VERSION : 0.1
   VAR_INPUT
      initValue : DWord;   // Initial value of CRC
      mask : DWord;   // Mask (CRC polynomial) / generator polynomial
      finalXorValue : DWord;   // Value to XOR the result with
      reflectInput : Bool;   // Reflect input (bits are used in reverse order)
      reflectResult : Bool;   // Reflect result (bits are used in reverse order)
   END_VAR
   VAR_IN_OUT
      inputArray : Array[*] of Byte;   // Input array / data stream
   END_VAR
   VAR_TEMP
      tempInput : Byte;   // Current input byte
      tempCRC : DWord;   // CRC checksum
      tempInvCRC : DWord;   // Inverted CRC checksum
      tempLowerLimit : DInt;   // Lower limit of input array
      tempUpperLimit : DInt;   // Upper limit of input array
      tempIndex1 : Int;   // -
      tempIndex2 : Int;   // -
   END_VAR
   // Ret_Val : CRC32 checksum
BEGIN
   //=============================================================================
   // Siemens AG
   // (c)Copyright 2017
   //-----------------------------------------------------------------------------
   // Library:       LGF (Library General Functions)
   // Tested with:   CPU1212C DC/DC/DC FW:V4.2
   // Engineering:   TIA Portal V14 SP1 Upd 5
   // Restrictions:  -
   // Requirements:  PLC (S7-1200 / S7-1500)
   // Functionality: CRC32
   //-----------------------------------------------------------------------------
   // Change log table:
   // Version  Date        In charge / Changes applied
   // 01.00.00 03.07.2018  Siemens Industry Online Support
   //                      First released version
   // 01.00.01 17.08.2018  Siemens Industry Online Support
   //                      Upgrade: TIA V15 Update 2
   // 01.00.02 23.11.2018  Siemens Industry Online Support
   //                      Upgrade: TIA V15.1
   //=============================================================================

   #tempLowerLimit := LOWER_BOUND(ARR := #inputArray, DIM := 1);
   #tempUpperLimit := UPPER_BOUND(ARR := #inputArray, DIM := 1);

   #tempCRC := #initValue;

   FOR #tempIndex1 := #tempLowerLimit TO #tempUpperLimit DO

     IF (#reflectInput = TRUE)
     THEN
       // Reverse bit order in input byte
       #tempInput.%X7 := #inputArray[#tempIndex1].%X0;
       #tempInput.%X6 := #inputArray[#tempIndex1].%X1;
       #tempInput.%X5 := #inputArray[#tempIndex1].%X2;
       #tempInput.%X4 := #inputArray[#tempIndex1].%X3;
       #tempInput.%X3 := #inputArray[#tempIndex1].%X4;
       #tempInput.%X2 := #inputArray[#tempIndex1].%X5;
       #tempInput.%X1 := #inputArray[#tempIndex1].%X6;
       #tempInput.%X0 := #inputArray[#tempIndex1].%X7;
     ELSE
       #tempInput := #inputArray[#tempIndex1];
     END_IF;

     #tempCRC := #tempCRC XOR SHL(IN := BYTE_TO_DWORD(#tempInput), N := 24);

     FOR #tempIndex2 := 0 TO 7 DO
       IF ((#tempCRC AND 16#80000000) <> 0)
       THEN
         #tempCRC := SHL(IN := #tempCRC, N := 1) XOR #mask;
       ELSE
         #tempCRC := SHL(IN := #tempCRC, N := 1);
       END_IF;
     END_FOR;

   END_FOR;

   IF (#reflectResult = TRUE)
   THEN
     // Reverse bit order in CRC checksum
     #tempInvCRC.%X31 := #tempCRC.%X0;
     #tempInvCRC.%X30 := #tempCRC.%X1;
     #tempInvCRC.%X29 := #tempCRC.%X2;
     #tempInvCRC.%X28 := #tempCRC.%X3;
     #tempInvCRC.%X27 := #tempCRC.%X4;
     #tempInvCRC.%X26 := #tempCRC.%X5;
     #tempInvCRC.%X25 := #tempCRC.%X6;
     #tempInvCRC.%X24 := #tempCRC.%X7;
     #tempInvCRC.%X23 := #tempCRC.%X8;
     #tempInvCRC.%X22 := #tempCRC.%X9;
     #tempInvCRC.%X21 := #tempCRC.%X10;
     #tempInvCRC.%X20 := #tempCRC.%X11;
     #tempInvCRC.%X19 := #tempCRC.%X12;
     #tempInvCRC.%X18 := #tempCRC.%X13;
     #tempInvCRC.%X17 := #tempCRC.%X14;
     #tempInvCRC.%X16 := #tempCRC.%X15;
     #tempInvCRC.%X15 := #tempCRC.%X16;
     #tempInvCRC.%X14 := #tempCRC.%X17;
     #tempInvCRC.%X13 := #tempCRC.%X18;
     #tempInvCRC.%X12 := #tempCRC.%X19;
     #tempInvCRC.%X11 := #tempCRC.%X20;
     #tempInvCRC.%X10 := #tempCRC.%X21;
     #tempInvCRC.%X9 := #tempCRC.%X22;
     #tempInvCRC.%X8 := #tempCRC.%X23;
     #tempInvCRC.%X7 := #tempCRC.%X24;
     #tempInvCRC.%X6 := #tempCRC.%X25;
     #tempInvCRC.%X5 := #tempCRC.%X26;
     #tempInvCRC.%X4 := #tempCRC.%X27;
     #tempInvCRC.%X3 := #tempCRC.%X28;
     #tempInvCRC.%X2 := #tempCRC.%X29;
     #tempInvCRC.%X1 := #tempCRC.%X30;
     #tempInvCRC.%X0 := #tempCRC.%X31;

     #LGF_CRC32 := #tempInvCRC XOR #finalXorValue;
   ELSE
     #LGF_CRC32 := #tempCRC XOR #finalXorValue;
   END_IF;
END_FUNCTION

// folder: Phisical_functions/LGF/6 Converter operations

FUNCTION "LGF_BinaryToGray" : DWord   // FC10021, SCL
{ S7_Optimized_Access := 'TRUE' }
   VAR_INPUT
      variableBinary : DWord;
   END_VAR
BEGIN
   //=============================================================================
   // SIEMENS AG
   // (c)Copyright 2017
   //-----------------------------------------------------------------------------
   // Library:       LGF(Library General Functions)
   // Tested with:   CPU1212C DC/DC/DC FW:V4.2
   // Engineering:   TIA Portal V14 Update 1
   // Restrictions:  -
   // Requirements:  PLC (S7-1200 / S7-1500)
   // Functionality: This function converts a binary value to a gray coded value
   //-----------------------------------------------------------------------------
   // Change log table:
   // Version  Date        In charge / Changes applied
   // 01.00.00 19.08.2015  Siemens Industry Online Support
   //                      First released version
   // 01.00.01 28.10.2015  Siemens Industry Online Support
   //                      Name changed
   // 01.00.02 02.01.2017  Siemens Industry Online Support
   //                      Upgrade: TIA Portal V14 Update 1
   // 01.00.03 17.08.2018  Siemens Industry Online Support
   //                      Upgrade: TIA V15 Update 2
   // 01.00.04 23.11.2018  Siemens Industry Online Support
   //                      Upgrade: TIA V15.1
   //=============================================================================

   #LGF_BinaryToGray := #variableBinary XOR SHR(IN := #variableBinary, N := 1);
END_FUNCTION

FUNCTION "LGF_GrayToBinary" : DWord   // FC10022, SCL
{ S7_Optimized_Access := 'TRUE' }
   VAR_INPUT
      variableGray : DWord;
   END_VAR
   VAR_TEMP
      tempBinaryBits : DWord;
   END_VAR
BEGIN
   //=============================================================================
   // SIEMENS AG
   // (c)Copyright 2017
   //-----------------------------------------------------------------------------
   // Library:       LGF(Library General Functions)
   // Tested with:   CPU1212C DC/DC/DC FW:V4.2
   // Engineering:   TIA Portal V14 Update 1
   // Restrictions:  -
   // Requirements:  PLC (S7-1200 / S7-1500)
   // Functionality: This function converts a gray coded value to a binary
   //-----------------------------------------------------------------------------
   // Change log table:
   // Version  Date        In charge / Changes applied
   // 01.00.00 19.08.2015  Siemens Industry Online Support
   //                      First released version
   // 01.00.01 28.10.2015  Siemens Industry Online Support
   //                      Name changed
   // 01.00.02 02.01.2017  Siemens Industry Online Support
   //                      Upgrade: TIA Portal V14 Update 1
   // 01.00.03 17.08.2018  Siemens Industry Online Support
   //                      Upgrade: TIA V15 Update 2
   // 01.00.04 23.11.2018  Siemens Industry Online Support
   //                      Upgrade: TIA V15.1
   //=============================================================================

   #tempBinaryBits := DW#16#0;

   #tempBinaryBits.%X31 := #variableGray.%X31;
   #tempBinaryBits.%X30 := #variableGray.%X30 XOR #tempBinaryBits.%X31;
   #tempBinaryBits.%X29 := #variableGray.%X29 XOR #tempBinaryBits.%X30;
   #tempBinaryBits.%X28 := #variableGray.%X28 XOR #tempBinaryBits.%X29;
   #tempBinaryBits.%X27 := #variableGray.%X27 XOR #tempBinaryBits.%X28;
   #tempBinaryBits.%X26 := #variableGray.%X26 XOR #tempBinaryBits.%X27;
   #tempBinaryBits.%X25 := #variableGray.%X25 XOR #tempBinaryBits.%X26;
   #tempBinaryBits.%X24 := #variableGray.%X24 XOR #tempBinaryBits.%X25;
   #tempBinaryBits.%X23 := #variableGray.%X23 XOR #tempBinaryBits.%X24;
   #tempBinaryBits.%X22 := #variableGray.%X22 XOR #tempBinaryBits.%X23;
   #tempBinaryBits.%X21 := #variableGray.%X21 XOR #tempBinaryBits.%X22;
   #tempBinaryBits.%X20 := #variableGray.%X20 XOR #tempBinaryBits.%X21;
   #tempBinaryBits.%X19 := #variableGray.%X19 XOR #tempBinaryBits.%X20;
   #tempBinaryBits.%X18 := #variableGray.%X18 XOR #tempBinaryBits.%X19;
   #tempBinaryBits.%X17 := #variableGray.%X17 XOR #tempBinaryBits.%X18;
   #tempBinaryBits.%X16 := #variableGray.%X16 XOR #tempBinaryBits.%X17;
   #tempBinaryBits.%X15 := #variableGray.%X15 XOR #tempBinaryBits.%X16;
   #tempBinaryBits.%X14 := #variableGray.%X14 XOR #tempBinaryBits.%X15;
   #tempBinaryBits.%X13 := #variableGray.%X13 XOR #tempBinaryBits.%X14;
   #tempBinaryBits.%X12 := #variableGray.%X12 XOR #tempBinaryBits.%X13;
   #tempBinaryBits.%X11 := #variableGray.%X11 XOR #tempBinaryBits.%X12;
   #tempBinaryBits.%X10 := #variableGray.%X10 XOR #tempBinaryBits.%X11;
   #tempBinaryBits.%X9 := #variableGray.%X9 XOR #tempBinaryBits.%X10;
   #tempBinaryBits.%X8 := #variableGray.%X8 XOR #tempBinaryBits.%X9;
   #tempBinaryBits.%X7 := #variableGray.%X7 XOR #tempBinaryBits.%X8;
   #tempBinaryBits.%X6 := #variableGray.%X6 XOR #tempBinaryBits.%X7;
   #tempBinaryBits.%X5 := #variableGray.%X5 XOR #tempBinaryBits.%X6;
   #tempBinaryBits.%X4 := #variableGray.%X4 XOR #tempBinaryBits.%X5;
   #tempBinaryBits.%X3 := #variableGray.%X3 XOR #tempBinaryBits.%X4;
   #tempBinaryBits.%X2 := #variableGray.%X2 XOR #tempBinaryBits.%X3;
   #tempBinaryBits.%X1 := #variableGray.%X1 XOR #tempBinaryBits.%X2;
   #tempBinaryBits.%X0 := #variableGray.%X0 XOR #tempBinaryBits.%X1;

   #LGF_GrayToBinary := #tempBinaryBits;
END_FUNCTION

FUNCTION "LGF_TemperatureConvert" : Real   // FC10023, SCL
{ S7_Optimized_Access := 'TRUE' }
   VAR_INPUT
      mode : Int;   // 1: Celsius in Fahrenheit, 2: Fahrenheit in Celsius, 3: Celsius in Kelvin, 4: Kelvin in Celsius, 5: Fahrenheit in Kelvin, 6: Kelvin in Fahrenheit
      temperature : Real;
   END_VAR
   VAR_OUTPUT
      error : Bool;
      status : Word;
   END_VAR
   VAR CONSTANT
      NO_ERROR : Word := 16#0000;
      NO_CURRENT_JOBS : Word := 16#7000;
      NO_MODE : Word := 16#8200;
   END_VAR
BEGIN
   //=============================================================================
   // SIEMENS AG
   // (c)Copyright 2017
   //-----------------------------------------------------------------------------
   // Library:       LGF (Library General Functions)
   // Tested with:   CPU1212C DC/DC/DC FW:V4.2
   // Engineering:   TIA Portal V14 Update 1
   // Restrictions:  -
   // Requirements:  PLC (S7-1200 / S7-1500)
   // Functionality: This function converts the temperature in another unit
   //-----------------------------------------------------------------------------
   // Change log table:
   // Version  Date        In charge / Changes applied
   // 01.00.00 19.08.2015  Siemens Industry Online Support
   //                      First released version
   // 01.00.01 02.01.2017  Siemens Industry Online Support
   //                      Upgrade: TIA Portal V14 Update 1
   // 01.00.02 17.08.2018  Siemens Industry Online Support
   //                      Upgrade: TIA V15 Update 2
   // 01.00.03 23.11.2018  Siemens Industry Online Support
   //                      Upgrade: TIA V15.1
   //=============================================================================

   //set "No current job" status
   #error := false;
   #status := #NO_CURRENT_JOBS;

   CASE #mode OF
       1:  // Celsius in Fahrenheit
          #LGF_TemperatureConvert := #temperature * 1.8 + 32.0; //F = C * 1.8 + 32
       2:  // Fahrenheit in Celsius
          #LGF_TemperatureConvert := (#temperature - 32.0)/ 1.8; //C = (F - 32) / 1.8
       3:  // Celsius in Kelvin
          #LGF_TemperatureConvert := #temperature + 273.15; //K = C + 273.15
       4:  // Kelvin in Celsius
          #LGF_TemperatureConvert := #temperature - 273.15; //C = K - 273.15
       5:  // Fahrenheit in Kelvin
          #LGF_TemperatureConvert := ((#temperature - 32.0) / 1.8) + 273.15 ; //K := ((C - 32.0) / 1.8) + 273.15
       6:  // Kelvin in Fahrenheit
          #LGF_TemperatureConvert := (#temperature - 273.15) * 1.8 + 32.0; //F := (K - 273.15) * 1.8 + 32.0
       ELSE  // no mode selected
         #error := true;
         #status:= #NO_MODE;
         #LGF_TemperatureConvert := 0.0;
         RETURN;
     END_CASE;

     #status := #NO_ERROR;
END_FUNCTION

FUNCTION "LGF_DTLtoString" : String   // FC10029, SCL
{ S7_Optimized_Access := 'TRUE' }
VERSION : 0.1
   VAR_INPUT
      inDTL : DTL;   // Date as DTL tag
      format : Bool;   // 1 = traditional, 0 = international
      separatorDate : Char;   // Separator between date components
   END_VAR
   VAR_TEMP
      tempString : String;   // -
      tempSepTime : Char;   // -
      tempSepTimeNano : Char;   // -
      tempPosYear : USInt;   // -
      tempPosMonth : USInt;   // -
      tempPosDay : USInt;   // -
      tempPosHour : USInt;   // -
      tempPosMinute : USInt;   // -
      tempPosSecond : USInt;   // -
      tempPosNanosecond : USInt;   // -
      tempPosSepYearMonth : USInt;   // -
      tempPosSepMonthDay : USInt;   // -
      tempPosSepHourMinute : USInt;   // -
      tempPosSepMinuteSecond : USInt;   // -
      tempPosSepSecondNanosecond : USInt;   // -
      tempCount : Int;   // -
   END_VAR
   // Ret_Val : Date as String tag
BEGIN
   //=============================================================================
   // Siemens AG
   // (c)Copyright 2017
   //-----------------------------------------------------------------------------
   // Library:       LGF (Library General Functions)
   // Tested with:   CPU1212C DC/DC/DC FW:V4.2
   // Engineering:   TIA Portal V14 Update 1
   // Restrictions:  -
   // Requirements:  PLC (S7-1200 / S7-1500)
   // Functionality: This function converts DTL into a string.  
   //-----------------------------------------------------------------------------
   // Change log table:
   // Version  Date        In charge / Changes applied
   // 01.00.00 15.06.2016  Siemens Industry Online Support
   //                      First released version
   // 01.00.01 02.01.2017  Siemens Industry Online Support
   //                      Upgrade: TIA Portal V14 Update 1
   // 01.00.02 17.08.2018  Siemens Industry Online Support
   //                      Upgrade: TIA V15 Update 2
   // 01.00.03 23.11.2018  Siemens Industry Online Support
   //                      Upgrade: TIA V15.1
   //=============================================================================

   // Initialization
   #tempString := '';
   #tempSepTime := ':';
   #tempSepTimeNano := '.';

   // Set format parameters for output string
   IF NOT #format
   THEN                                          // International ISO 8601
     #tempPosYear := 1;                          // DTL  | Y| Y| Y| Y| -| M| M| -| D| D|  | H| H| :| M| M| :| S| S| .|NS|NS|NS|NS|NS|NS|NS|NS|NS
     #tempPosMonth := 6;                         // -----|--|--|--|--|--|--|--|--|--|--|--|--|--|--|--|--|--|--|--|--|--|--|--|--|--|--|--|--|--
     #tempPosDay := 9;                           // Pos  | 1| 2| 3| 4| 5| 6| 7| 8| 9|10|11|12|13|14|15|16|17|18|19|20|21|22|23|24|25|26|27|28|29
     #tempPosHour := 12;
     #tempPosMinute := 15;
     #tempPosSecond := 18;
     #tempPosNanosecond := 21;
     #tempPosSepYearMonth := 5;
     #tempPosSepMonthDay := 8;
     #tempPosSepHourMinute := 14;
     #tempPosSepMinuteSecond := 17;
     #tempPosSepSecondNanosecond := 20;
   ELSE                                          // Traditional (EU)
     #tempPosYear := 7;                          // DTL  | D| D| -| M| M| -| Y| Y| Y| Y|  | H| H| :| M| M| :| S| S| .|NS|NS|NS|NS|NS|NS|NS|NS|NS
     #tempPosMonth := 4;                         // -----|--|--|--|--|--|--|--|--|--|--|--|--|--|--|--|--|--|--|--|--|--|--|--|--|--|--|--|--|--
     #tempPosDay := 1;                           // Pos  | 1| 2| 3| 4| 5| 6| 7| 8| 9|10|11|12|13|14|15|16|17|18|19|20|21|22|23|24|25|26|27|28|29
     #tempPosHour := 12;
     #tempPosMinute := 15;
     #tempPosSecond := 18;
     #tempPosNanosecond := 21;
     #tempPosSepYearMonth := 6;
     #tempPosSepMonthDay := 3;
     #tempPosSepHourMinute := 14;
     #tempPosSepMinuteSecond := 17;
     #tempPosSepSecondNanosecond := 20;
   END_IF;

   // Convert "Value" into "String" and place at the right position
   VAL_STRG(FORMAT := W#16#0000,
            IN := #inDTL.YEAR,
            P := #tempPosYear,
            PREC := 0,
            SIZE := 4,
            OUT => #tempString);    // DTL YEAR --> String --> #tempPosYear

   VAL_STRG(FORMAT := W#16#0000,
            IN := #inDTL.MONTH,
            P := #tempPosMonth,
            PREC := 0,
            SIZE := 2,
            OUT => #tempString);     // DTL MONTH --> String --> #tempPosMonth

   VAL_STRG(FORMAT := W#16#0000,
            IN := #inDTL.DAY,
            P := #tempPosDay,
            PREC := 0,
            SIZE := 2,
            OUT => #tempString);     // DTL DAY --> String --> #tempPosDay

   VAL_STRG(FORMAT := W#16#0000,
            IN := #inDTL.HOUR,
            P := #tempPosHour,
            PREC := 0,
            SIZE := 2,
            OUT => #tempString);     // DTL HOUR --> String --> #tempPosHour

   VAL_STRG(FORMAT := W#16#0000,
            IN := #inDTL.MINUTE,
            P := #tempPosMinute,
            PREC := 0,
            SIZE := 2,
            OUT => #tempString);     // DTL MINUTE --> String --> #tempPosMinute

   VAL_STRG(FORMAT := W#16#0000,
            IN := #inDTL.SECOND,
            P := #tempPosSecond,
            PREC := 0,
            SIZE := 2,
            OUT => #tempString);     // DTL SECOND --> String --> #tempPosSecond

   VAL_STRG(FORMAT := W#16#0000,
            IN := #inDTL.NANOSECOND,
            P := #tempPosNanosecond,
            PREC := 0,
            SIZE := 9,
            OUT => #tempString);     // DTL NANOSECOND --> String --> #tempPosNanosecond

   // Place separators at the right position in the string
   #tempString[#tempPosSepYearMonth] := #separatorDate;
   #tempString[#tempPosSepMonthDay] := #separatorDate;
   #tempString[#tempPosSepHourMinute] := #tempSepTime;
   #tempString[#tempPosSepMinuteSecond] := #tempSepTime;
   #tempString[#tempPosSepSecondNanosecond] := #tempSepTimeNano;

   // Correcting the string, due to the conversion of a leading "0" value into a "blank".
   // Replacing of "blank" by "0"
   IF (#tempString[#tempPosMonth] = ' ')
   THEN
     #tempString[#tempPosMonth] := '0';
   END_IF;

   IF (#tempString[#tempPosDay] = ' ')
   THEN
     #tempString[#tempPosDay] := '0';
   END_IF;

   IF (#tempString[#tempPosHour] = ' ')
   THEN
     #tempString[#tempPosHour] := '0';
   END_IF;

   IF (#tempString[#tempPosMinute] = ' ')
   THEN
     #tempString[#tempPosMinute] := '0';
   END_IF;

   IF (#tempString[#tempPosSecond] = ' ')
   THEN
     #tempString[#tempPosSecond] := '0';
   END_IF;

   FOR #tempCount := 0 TO 5 BY 1
   DO
     IF (#tempString[#tempPosNanosecond + #tempCount] = ' ')
     THEN
       #tempString[#tempPosNanosecond + #tempCount] := '0';
     ELSE
       EXIT;
     END_IF;
   END_FOR;

   #LGF_DTLtoString := #tempString;
END_FUNCTION

FUNCTION "LGF_StringToDTL" : DTL   // FC10030, SCL
{ S7_Optimized_Access := 'TRUE' }
VERSION : 0.1
   VAR_INPUT
      inString : String;   // Date as String tag
      format : Bool;   // Format of inString/ 0=traditional; 1=international
   END_VAR
   VAR_OUTPUT
      error : Bool;   // "0" = no error; "1" = error
      status : Word;   // status and error codes
   END_VAR
   VAR_TEMP
      tempCounter : Int;   // -
      tempOutput : DTL;   // -
      tempYear : String;   // -
      tempMonth : String;   // -
      tempDay : String;   // -
      tempHour : String;   // -
      tempMinute : String;   // -
      tempSecond : String;   // -
      tempNanosecond : String;   // -
      tempPosYear : USInt;   // -
      tempPosMonth : USInt;   // -
      tempPosDay : USInt;   // -
      tempPosHour : USInt;   // -
      tempPosMinute : USInt;   // -
      tempPosSecond : USInt;   // -
      tempPosNanosecond : USInt;   // -
      tempPosSepYearMonth : USInt;   // -
      tempPosSepMonthDay : USInt;   // -
      tempPosSepHourMinute : USInt;   // -
      tempPosSepMinuteSecond : USInt;   // -
      tempPosSepSecondNanosecond : USInt;   // -
   END_VAR
   // Ret_Val : Date as DTL tag / -
   VAR CONSTANT
      NO_ERROR : Word := 16#0000;   // -
      NO_CURRENT_JOBS : Word := 16#7000;   // -
      ERROR_FORMAT_YEAR : Word := 16#8201;   // -
      ERROR_FORMAT_MONTH : Word := 16#8202;   // -
      ERROR_FORMAT_DAY : Word := 16#8203;   // -
      ERROR_FORMAT_HOUR : Word := 16#8204;   // -
      ERROR_FORMAT_MINUTE : Word := 16#8205;   // -
      ERROR_FORMAT_SECOND : Word := 16#8206;   // -
      ERROR_FORMAT_NANOSECOND : Word := 16#8207;   // -
      INITIAL_VALUE : DTL := DTL#1970-01-01-00:00:00.0;   // -
   END_VAR
BEGIN
   //=============================================================================
   // SIEMENS AG
   // (c)Copyright 2017
   //-----------------------------------------------------------------------------
   // Library:       LGF (Library General Functions)
   // Tested with:   CPU1212C DC/DC/DC FW:V4.2
   // Engineering:   TIA Portal V14 Update 1
   // Restrictions:  -
   // Requirements:  PLC (S7-1200 / S7-1500)
   // Functionality: This function converts a string including date and time  
   //                information into DTL format.
   //-----------------------------------------------------------------------------
   // Change log table:
   // Version  Date        In charge / Changes applied
   // 01.00.00 15.06.2016  Siemens Industry Online Support
   //                      First released version
   // 01.00.01 02.01.2017  Siemens Industry Online Support
   //                      Upgrade: TIA Portal V14 Update 1
   // 01.00.02 17.08.2018  Siemens Industry Online Support
   //                      Upgrade: TIA V15 Update 2
   // 01.00.03 23.11.2018  Siemens Industry Online Support
   //                      Upgrade: TIA V15.1
   //-----------------------------------------------------------------------------
   //Status Codes:
   // 16#0000:  No errors
   // 16#7000:  Initial state
   // 16#820x:  Wrong format of the input string (Note position of components in
   //           the string)
   //=============================================================================

   //Set initial parameters
   #error := FALSE;
   #status := #NO_ERROR;

   IF #inString = ''
   THEN
     #LGF_StringToDTL := #INITIAL_VALUE;
     #status := #NO_CURRENT_JOBS;
     RETURN;
   END_IF;

   // Set format parameters for input string
   IF NOT #format
   THEN
     #tempPosYear := 1;                          // DTL  | Y| Y| Y| Y| -| M| M| -| D| D|  | H| H| :| M| M| :| S| S| .|NS|NS|NS|NS|NS|NS|NS|NS|NS
     #tempPosMonth := 6;                         // -----|--|--|--|--|--|--|--|--|--|--|--|--|--|--|--|--|--|--|--|--|--|--|--|--|--|--|--|--|--
     #tempPosDay := 9;                           // Pos  | 1| 2| 3| 4| 5| 6| 7| 8| 9|10|11|12|13|14|15|16|17|18|19|20|21|22|23|24|25|26|27|28|29
     #tempPosHour := 12;
     #tempPosMinute := 15;
     #tempPosSecond := 18;
     #tempPosNanosecond := 21;
     #tempPosSepYearMonth := 5;
     #tempPosSepMonthDay := 8;
     #tempPosSepHourMinute := 14;
     #tempPosSepMinuteSecond := 17;
     #tempPosSepSecondNanosecond := 20;
   ELSE
     #tempPosYear := 7;                          // DTL  | D| D| -| M| M| -| Y| Y| Y| Y|  | H| H| :| M| M| :| S| S| .|NS|NS|NS|NS|NS|NS|NS|NS|NS
     #tempPosMonth := 4;                         // -----|--|--|--|--|--|--|--|--|--|--|--|--|--|--|--|--|--|--|--|--|--|--|--|--|--|--|--|--|--
     #tempPosDay := 1;                           // Pos  | 1| 2| 3| 4| 5| 6| 7| 8| 9|10|11|12|13|14|15|16|17|18|19|20|21|22|23|24|25|26|27|28|29
     #tempPosHour := 12;
     #tempPosMinute := 15;
     #tempPosSecond := 18;
     #tempPosNanosecond := 21;
     #tempPosSepYearMonth := 6;
     #tempPosSepMonthDay := 3;
     #tempPosSepHourMinute := 14;
     #tempPosSepMinuteSecond := 17;
     #tempPosSepSecondNanosecond := 20;
   END_IF;

   // Separating the input string into components of DTL
   #tempYear := MID(IN := #inString, L := 4, P := #tempPosYear);
   #tempMonth := MID(IN := #inString, L := 2, P := #tempPosMonth);
   #tempDay := MID(IN := #inString, L := 2, P := #tempPosDay);
   #tempHour := MID(IN := #inString, L := 2, P := #tempPosHour);
   #tempMinute := MID(IN := #inString, L := 2, P := #tempPosMinute);
   #tempSecond := MID(IN := #inString, L := 2, P := #tempPosSecond);
   #tempNanosecond := MID(IN := #inString, L := 9, P := #tempPosNanosecond);

   // Replacing of the "blan" in the nanosecondstring by "0"
   // Effect:   xx.1 --> xx.1 AND NOT xx.1 --> xx.000000001
   FOR #tempCounter := 1 TO 9 BY 1
   DO
     IF #tempNanosecond[#tempCounter] = ' '
     THEN
       #tempNanosecond[#tempCounter] := '0';
     END_IF;
   END_FOR;

   // Converting separated String components into DTL values
   STRG_VAL(FORMAT := W#16#0000,
            IN := #tempYear,
            OUT => #tempOutput.YEAR,
            P := 1);

   STRG_VAL(FORMAT := W#16#0000,
            IN := #tempMonth,
            OUT => #tempOutput.MONTH,
            P := 1);

   STRG_VAL(FORMAT := W#16#0000,
            IN := #tempDay,
            OUT => #tempOutput.DAY,
            P := 1);

   STRG_VAL(FORMAT := W#16#0000,
            IN := #tempHour,
            OUT => #tempOutput.HOUR,
            P := 1);

   STRG_VAL(FORMAT := W#16#0000,
            IN := #tempMinute,
            OUT => #tempOutput.MINUTE,
            P := 1);

   STRG_VAL(FORMAT := W#16#0000,
            IN := #tempSecond,
            OUT => #tempOutput.SECOND,
            P := 1);

   STRG_VAL(FORMAT := W#16#0000,
            IN := #tempNanosecond,
            OUT => #tempOutput.NANOSECOND,
            P := 1);

   // Format check
   IF (#tempOutput.YEAR < 1970) OR (2262 < #tempOutput.YEAR)
   THEN
     #error := TRUE;
     #status := #ERROR_FORMAT_YEAR;
     #LGF_StringToDTL := #INITIAL_VALUE;
     RETURN;
   END_IF;

   IF (#tempOutput.MONTH < 1) OR (12 < #tempOutput.MONTH)
   THEN
     #error := TRUE;
     #status := #ERROR_FORMAT_MONTH;
     #LGF_StringToDTL := #INITIAL_VALUE;
     RETURN;
   END_IF;

   IF (#tempOutput.DAY < 1) OR (31 < #tempOutput.DAY)
   THEN
     #error := TRUE;
     #status := #ERROR_FORMAT_DAY;
     #LGF_StringToDTL := #INITIAL_VALUE;
     RETURN;
   END_IF;

   IF (#tempOutput.HOUR < 0) OR (23 < #tempOutput.HOUR)
   THEN
     #error := TRUE;
     #status := #ERROR_FORMAT_HOUR;
     #LGF_StringToDTL := #INITIAL_VALUE;
     RETURN;
   END_IF;

   IF (#tempOutput.MINUTE < 0) OR (59 < #tempOutput.MINUTE)
   THEN
     #error := TRUE;
     #status := #ERROR_FORMAT_MINUTE;
     #LGF_StringToDTL := #INITIAL_VALUE;
     RETURN;
   END_IF;

   IF (#tempOutput.SECOND < 0) OR (59 < #tempOutput.SECOND)
   THEN
     #error := TRUE;
     #status := #ERROR_FORMAT_SECOND;
     #LGF_StringToDTL := #INITIAL_VALUE;
     RETURN;
   END_IF;

   IF (#tempOutput.NANOSECOND < 0) OR (999999999 < #tempOutput.NANOSECOND)
   THEN
     #error := TRUE;
     #status := #ERROR_FORMAT_NANOSECOND;
     #LGF_StringToDTL := #INITIAL_VALUE;
     RETURN;
   END_IF;

   #LGF_StringToDTL := #tempOutput;
END_FUNCTION

FUNCTION "LGF_ScaleLinear" : Void   // FC10039, SCL
{ S7_Optimized_Access := 'TRUE' }
VERSION : 0.1
   VAR_INPUT
      x : LReal;   // Value to be scaled
      x1 : LReal;   // x coordinate for point 1
      y1 : LReal;   // y coordinate for point 1
      x2 : LReal;   // x coordinate for point 2
      y2 : LReal;   // y coordinate for point 2
      yMin : LReal;   // Lower limit for the output value
      yMax : LReal;   // Upper limit for the output value
   END_VAR
   VAR_OUTPUT
      y : LReal;   // Scaled value y
      error : Bool;   // FALSE: No error / TRUE: Error.
      status : Word;   // Error information.
   END_VAR
   VAR_TEMP
      tempY : LReal;   // Temporary scaled value y
   END_VAR
   // Ret_Val : -
   VAR CONSTANT
      NO_ERROR : Word := 16#0000;   // No error
      "LOW_LIM_OVER UP_LIM" : Word := 16#8204;   // Lower limit is greater than upper limit
      Y_LIMITED_TO_YMIN : Word := 16#8205;   // Y value limited to yMin
      Y_LIMITED_TO_YMAX : Word := 16#8206;   // Y value limited to yMax
   END_VAR
BEGIN
   //=============================================================================
   // Siemens AG
   // (c)Copyright 2017
   //-----------------------------------------------------------------------------
   // Library:       LGF (Library General Functions)
   // Tested with:   CPU1212C DC/DC/DC FW:V4.2
   // Engineering:   TIA Portal V14 Upd 1
   // Restrictions:  -
   // Requirements:  PLC (S7-1200 / S7-1500)
   // Functionality: This function scales a value (INT/REAL)
   //-----------------------------------------------------------------------------
   // Change log table:
   // Version  Date        In charge / Changes applied
   // 01.00.00 27.01.2017  Siemens Industry Online Support
   //                      First released version
   // 01.00.01 17.08.2018  Siemens Industry Online Support
   //                      Upgrade: TIA V15 Update 2
   // 01.00.02 23.11.2018  Siemens Industry Online Support
   //                      Upgrade: TIA V15.1
   // 02.00.00 25.01.2019  Siemens Industry Online Support
   //                      Data type changed from Variant to LReal
   //-----------------------------------------------------------------------------
   //Status Codes: 16#0000 - no error
   //              16#8204 - Lower limit is greater than upper limit. 
   //=============================================================================

   #error := FALSE;
   #status := #NO_ERROR;

   IF (#yMin > #yMax)
   THEN
     #error := TRUE;
     #status := #"LOW_LIM_OVER UP_LIM";
     RETURN;
   END_IF;

   // Scale algorithm
   IF ((#x2 - #x1) = 0.0)
   THEN
     #tempY := #y1;
   ELSE
     #tempY := (#y2 - #y1) / (#x2 - #x1) * (#x - #x1) + #y1;
   END_IF;

   // Check upper and lower limits
   IF (#tempY < #yMin)
   THEN
     #y := #yMin;
     #status := #Y_LIMITED_TO_YMIN;  //No error, only for information
   ELSIF (#tempY > #yMax)
   THEN
     #y := #yMax;
     #status := #Y_LIMITED_TO_YMAX;  //No error, only for information
   ELSE
     #y := #tempY;
   END_IF;
END_FUNCTION

FUNCTION "LGF_StringToTaddr" : TADDR_Param   // FC10041, SCL
{ S7_Optimized_Access := 'TRUE' }
VERSION : 0.1
   VAR_INPUT
      ipAddressString : String;   // in the format of '192.168.1.200:55047' Port number is optional [ you can obmit the : and following port number]
   END_VAR
   VAR_OUTPUT
      error : Bool;   // "0" = no error; "1" = error
      status : Word;   // status and error codes
   END_VAR
   VAR_TEMP
      tempCharPosition : Int;
      tempAddressString : String;
      tempOctetString : String[4];
      tempUInt : UInt;
      tempPortNumberIsSpecified : Bool;
      tempIpAdressTaddr : TADDR_Param;
   END_VAR
   VAR CONSTANT
      NO_ERROR : Word := 16#0000;   // Status no error
      WRONG_VALUE_POS1 : Word := 16#8101;   // Wrong value on position 1
      WRONG_VALUE_POS2 : Word := 16#8102;   // Wrong value on position 2
      WRONG_VALUE_POS3 : Word := 16#8103;   // Wrong value on position 3
      WRONG_VALUE_POS4 : Word := 16#8104;   // Wrong value on position 4
      WRONG_VALUE_PORT : Word := 16#8105;   // Wrong value on port position
      MAX_USINT : USInt := 255;
      MAX_UINT : UInt := 65535;
      EMPTY_STRING : String := '';
      MAX_CHAR_FOR_IP_PART : Int := 4;
      MAX_CHAR_FOR_PORT_PART : Int := 5;
      INIT_VAL : USInt := 0;
      NO_POS : Int := 0;
   END_VAR
BEGIN
   //=============================================================================
   // SIEMENS AG
   // (c)Copyright 2017
   //-----------------------------------------------------------------------------
   // Library:       LGF (Library General Functions)
   // Tested with:   CPU1212C DC/DC/DC FW:V4.2
   // Engineering:   TIA Portal V14 Upd 1
   // Restrictions:  -
   // Requirements:  PLC (S7-1200 / S7-1500)
   // Functionality: This function converts a string IP Address
   //                into TADDR Param format.
   //-----------------------------------------------------------------------------
   // Change log table:
   // Version  Date        In charge Changes applied
   // 01.00.00 30.01.2017  Siemens Industry Online Support
   //                      First released version
   // 01.00.01 17.08.2018  Siemens Industry Online Support
   //                      Upgrade: TIA V15 Update 2
   // 01.00.02 23.11.2018  Siemens Industry Online Support
   //                      Upgrade: TIA V15.1
   //-----------------------------------------------------------------------------
   //Status Codes:
   // 16#0000:  No errors
   // 16#8101:  Wrong value on position 1
   // 16#8102:  Wrong value on position 2
   // 16#8103:  Wrong value on position 3
   // 16#8104:  Wrong value on position 4
   // 16#8105:  Wrong value on port position
   //=============================================================================

   // Initialization
   #error := FALSE;
   #status := #NO_ERROR;
   #tempAddressString := #ipAddressString;
   #LGF_StringToTaddr.REM_IP_ADDR[1] := #INIT_VAL;
   #LGF_StringToTaddr.REM_IP_ADDR[2] := #INIT_VAL;
   #LGF_StringToTaddr.REM_IP_ADDR[3] := #INIT_VAL;
   #LGF_StringToTaddr.REM_IP_ADDR[4] := #INIT_VAL;
   #LGF_StringToTaddr.REM_PORT_NR := #INIT_VAL;

   // Process the 1st octet of the IP Address
   #tempCharPosition := FIND(IN1 := #tempAddressString, IN2 := '.');
   IF #tempCharPosition > #MAX_CHAR_FOR_IP_PART THEN
     #error := TRUE;
     #status := #WRONG_VALUE_POS1;
     RETURN;
   ELSE
     #tempOctetString := LEFT(IN := #tempAddressString, L := #tempCharPosition - 1);
     // Check if string is empty
     IF #tempOctetString = #EMPTY_STRING THEN
       #error := TRUE;
       #status := #WRONG_VALUE_POS1;
       RETURN;
     ELSE
       #tempAddressString := DELETE(IN := #tempAddressString, P := 1, L := #tempCharPosition);
     END_IF;
   END_IF;

   // Convert the 1st octet string to numerical value
   STRG_VAL(IN := #tempOctetString,
            FORMAT := W#16#0000,
            P := 1,
            OUT => #tempUInt);

     IF #tempUInt > #MAX_USINT THEN
       #error := TRUE;
       #status := #WRONG_VALUE_POS1;
       RETURN;
     ELSE
       #tempIpAdressTaddr.REM_IP_ADDR[1] := UINT_TO_BYTE(#tempUInt);
     END_IF;


   // Process the 2nd octetstring of the IP Address
   #tempCharPosition := FIND(IN1 := #tempAddressString, IN2 := '.');
   IF #tempCharPosition > #MAX_CHAR_FOR_IP_PART THEN
     #error := TRUE;
     #status := #WRONG_VALUE_POS2;
     RETURN;
   ELSE
     #tempOctetString := LEFT(IN := #tempAddressString, L := #tempCharPosition - 1);
     IF #tempOctetString = #EMPTY_STRING THEN
       #error := TRUE;
       #status := #WRONG_VALUE_POS2;
       RETURN;
     ELSE
       #tempAddressString := DELETE(IN := #tempAddressString, P := 1, L := #tempCharPosition);
     END_IF;
   END_IF;

   // Convert the 2nd octet string TO numerical value
   STRG_VAL(IN := #tempOctetString,
            FORMAT := W#16#0000,
            P := 1,
            OUT => #tempUInt);

   IF #tempUInt > #MAX_USINT THEN
     #error := TRUE;
     #status := #WRONG_VALUE_POS2;
     RETURN;
   ELSE
     #tempIpAdressTaddr.REM_IP_ADDR[2] := UINT_TO_BYTE(#tempUInt);
   END_IF;

   // Process the 3rd octet of the IP Address
   #tempCharPosition := FIND(IN1 := #tempAddressString, IN2 := '.');
   IF #tempCharPosition > #MAX_CHAR_FOR_IP_PART THEN
     #error := TRUE;
     #status := #WRONG_VALUE_POS3;
     RETURN;
   ELSE
     #tempOctetString := LEFT(IN := #tempAddressString, L := #tempCharPosition - 1);
     // Check if string is empty
     IF #tempOctetString = #EMPTY_STRING THEN
       #error := TRUE;
       #status := #WRONG_VALUE_POS3;
       RETURN;
     ELSE
       #tempAddressString := DELETE(IN := #tempAddressString, P := 1, L := #tempCharPosition);
     END_IF;
   END_IF;

   //Convert the 3rd octet string to numerical value
   STRG_VAL(IN := #tempOctetString,
            FORMAT := W#16#0000,
            P := 1,
            OUT => #tempUInt);
   IF #tempUInt > #MAX_USINT
   THEN
     #error := TRUE;
     #status := #WRONG_VALUE_POS3;
     RETURN;
   ELSE
     #tempIpAdressTaddr.REM_IP_ADDR[3] := UINT_TO_BYTE(#tempUInt);
   END_IF;

   // Process the 4th octet of the IP Address
   #tempCharPosition := FIND(IN1 := #tempAddressString, IN2 := '.');
   IF #tempCharPosition > #NO_POS THEN
     #error := TRUE;
     #status := #WRONG_VALUE_POS4;
     RETURN;
   ELSE
     #tempCharPosition := FIND(IN1 := #tempAddressString, IN2 := ':');
   END_IF;

   // Check if Port number added
   #tempPortNumberIsSpecified := (#tempCharPosition > #NO_POS);
   IF #tempCharPosition > #MAX_CHAR_FOR_PORT_PART THEN
     #error := TRUE;
     #status := #WRONG_VALUE_PORT;
     RETURN;
   END_IF;
   IF NOT #tempPortNumberIsSpecified THEN
     #tempCharPosition := LEN(#tempAddressString) + 1;
   END_IF;

   #tempOctetString := LEFT(IN := #tempAddressString, L := #tempCharPosition - 1);
   // Check if string is empty
   IF #tempOctetString = #EMPTY_STRING THEN
     #error := TRUE;
     #status := #WRONG_VALUE_POS4;
     RETURN;
   ELSE
     #tempAddressString := DELETE(IN := #tempAddressString, P := 1, L := #tempCharPosition);
   END_IF;

   // Convert the 4th octet string to numerical value
   STRG_VAL(IN := #tempOctetString,
            FORMAT := W#16#0000,
            P := 1,
            OUT => #tempUInt);

   IF #tempUInt > #MAX_USINT THEN
     #error := TRUE;
     #status := #WRONG_VALUE_POS4;
     RETURN;
   ELSE
     #tempIpAdressTaddr.REM_IP_ADDR[4] := UINT_TO_BYTE(#tempUInt);
   END_IF;

   // If the string contains a port number too, parse it
   IF #tempPortNumberIsSpecified THEN
     // Convert the port number string to numerical value
     STRG_VAL(IN := #tempAddressString,
              FORMAT := W#16#0000,
              P := 1,
              OUT => #tempUInt);
     IF #tempUInt > #MAX_UINT OR #tempUInt = 0 THEN
       #error := TRUE;
       #status := #WRONG_VALUE_PORT;
       RETURN;
     ELSE
       #tempIpAdressTaddr.REM_PORT_NR := #tempUInt;
     END_IF;
   END_IF;

   // Write Outputs
   #LGF_StringToTaddr := #tempIpAdressTaddr;
END_FUNCTION

FUNCTION "LGF_TaddrToString" : String   // FC10042, SCL
{ S7_Optimized_Access := 'TRUE' }
VERSION : 0.1
   VAR_INPUT
      ipAdressTaddr : TADDR_Param;
   END_VAR
   VAR_TEMP
      tempIpAddressString : String;
      tempSpaceLocation : Int;
   END_VAR
BEGIN
   //=============================================================================
   // SIEMENS AG
   // (c)Copyright 2017
   //-----------------------------------------------------------------------------
   // Library:       LGF (Library General Functions)
   // Tested with:   CPU1212C DC/DC/DC FW:V4.2
   // Engineering:   TIA Portal V14 Upd 1
   // Restrictions:  -
   // Requirements:  PLC (S7-1200 / S7-1500)
   // Functionality: This function converts  TADDR Param into a string IP Address
   //                format.
   //-----------------------------------------------------------------------------
   // Change log table:
   // Version  Date        In charge /Changes applied
   // 01.00.00 19.01.2017  Siemens Industry Online Support
   //                      First released version
   // 01.00.01 17.08.2018  Siemens Industry Online Support
   //                      Upgrade: TIA V15 Update 2
   // 01.00.02 23.11.2018  Siemens Industry Online Support
   //                      Upgrade: TIA V15.1
   //=============================================================================

   // Convert the first IPV4 Octet to a string
   VAL_STRG(IN := #ipAdressTaddr.REM_IP_ADDR[1],
            SIZE := 3,
            PREC := 0,
            FORMAT := 0,
            P := 1,
            OUT => #tempIpAddressString);

   #tempIpAddressString[4] := '.';

   // Convert the second IPV4 Octet to a string
   VAL_STRG(IN := #ipAdressTaddr.REM_IP_ADDR[2],
            SIZE := 3,
            PREC := 0,
            FORMAT := 0,
            P := 5,
            OUT => #tempIpAddressString);

   #tempIpAddressString[8] := '.';

   // Convert the third IPV4 Octet to a string
   VAL_STRG(IN := #ipAdressTaddr.REM_IP_ADDR[3],
            SIZE := 3,
            PREC := 0,
            FORMAT := 0,
            P := 9,
            OUT => #tempIpAddressString);

   #tempIpAddressString[12] := '.';

   // Convert the fourth IPV4 Octet to a string
   VAL_STRG(IN := #ipAdressTaddr.REM_IP_ADDR[4],
            SIZE := 3,
            PREC := 0,
            FORMAT := 0,
            P := 13,
            OUT => #tempIpAddressString);

   // If the Port number is specified, copy it to the string following the ':' seperator
   IF #ipAdressTaddr.REM_PORT_NR > 0 THEN
     #tempIpAddressString[16] := ':';
     //Convert the port number to a string
     VAL_STRG(IN := #ipAdressTaddr.REM_PORT_NR,
              SIZE := 5,
              PREC := 0,
              FORMAT := 0,
              P := 17,
              OUT => #tempIpAddressString);
   END_IF;

   // Delete all spaces in the string
   #tempSpaceLocation := 1;

   WHILE #tempSpaceLocation > 0 DO
     #tempSpaceLocation := FIND(IN1 := #tempIpAddressString, IN2 := ' ');
     IF #tempSpaceLocation > 0 THEN
       #tempIpAddressString := DELETE(IN := #tempIpAddressString, L := 1, P := #tempSpaceLocation);
     END_IF;
   END_WHILE;

   // Write outputs
   #LGF_TaddrToString := #tempIpAddressString;
END_FUNCTION

FUNCTION "LGF_TimeToString" : String   // FC10043, SCL
{ S7_Optimized_Access := 'TRUE' }
VERSION : 0.1
   VAR_INPUT
      timeValue : Time;   // Time value to convert
   END_VAR
   VAR_OUTPUT
      stringDay : String;   // String for day
      stringHour : String;   // String for hour
      stringMinute : String;   // String for minute
      stringSecond : String;   // String for second
      stringMilliSecond : String;   // String for millisecond
   END_VAR
   VAR_TEMP
      tempStringTime : String;
      tempTimeInt : DInt;
      tempModDays : DInt;
      tempModHours : DInt;
      tempModMinutes : DInt;
      tempModSecond : DInt;
      tempModMilliSecond : DInt;
      tempDivDays : DInt;
      tempDivHours : DInt;
      tempDivMinutes : DInt;
      tempDivSecond : DInt;
      tempDivMillisecond : DInt;
   END_VAR
   VAR CONSTANT
      MS_PER_DAY : DInt := 86400000;
      MS_PER_HOUR : DInt := 3600000;
      MS_PER_MINUTE : DInt := 60000;
      MS_PER_SECOND : DInt := 1000;
   END_VAR
BEGIN
   //=============================================================================
   // Siemens AG
   // (c)Copyright 2017
   //-----------------------------------------------------------------------------
   // Library:       LGF (Library General Functions)
   // Tested with:   CPU1212C DC/DC/DC FW:V4.2
   // Engineering:   TIA Portal V14 SP1 Upd 5
   // Restrictions:  -
   // Requirements:  PLC (S7-1200 / S7-1500)
   // Functionality: This function converts a time value to a string
   //-----------------------------------------------------------------------------
   // Change log table:
   // Version  Date        In charge / Changes applied
   // 01.00.00 03.07.2018  Siemens Industry Online Support
   //                      First released version
   // 01.00.01 17.08.2018  Siemens Industry Online Support
   //                      Upgrade: TIA V15 Update 2
   // 01.00.02 23.11.2018  Siemens Industry Online Support
   //                      Upgrade: TIA V15.1
   //=============================================================================

   // Init string
   #tempStringTime := '0';

   #tempTimeInt := TIME_TO_DINT(#timeValue);

   #tempDivDays := #tempTimeInt / #MS_PER_DAY;
   #tempModDays := #tempTimeInt MOD #MS_PER_DAY;

   #tempDivHours := #tempModDays / #MS_PER_HOUR;
   #tempModHours := #tempModDays MOD #MS_PER_HOUR;

   #tempDivMinutes := #tempModHours / #MS_PER_MINUTE;
   #tempModMinutes := #tempModHours MOD #MS_PER_MINUTE;

   #tempDivSecond := #tempModMinutes / #MS_PER_SECOND;
   #tempModSecond := #tempModMinutes MOD #MS_PER_SECOND;

   #tempDivMillisecond := #tempModSecond;


   #stringDay := DELETE(IN := DINT_TO_STRING(#tempDivDays), L := 1, P := 1);
   #stringHour := DELETE(IN := DINT_TO_STRING(#tempDivHours), L := 1, P := 1);;
   #stringMinute := DELETE(IN := DINT_TO_STRING(#tempDivMinutes), L := 1, P := 1);
   #stringSecond := DELETE(IN := DINT_TO_STRING(#tempDivSecond), L := 1, P := 1);
   #stringMilliSecond := DELETE(IN := DINT_TO_STRING(#tempDivMillisecond), L := 1, P := 1);

   IF (#tempDivMillisecond > 0)
   THEN
     #tempStringTime := CONCAT(IN1 := #stringMilliSecond, IN2 := 'MS');
   END_IF;

   IF (#tempDivSecond > 0)
   THEN
     #tempStringTime := CONCAT(IN1 := #stringSecond, IN2 := 'S', IN3 := #stringMilliSecond, IN4 := 'MS');
   END_IF;

   IF (#tempDivMinutes > 0)
   THEN
     #tempStringTime := CONCAT(IN1 := #stringMinute, IN2 := 'M', IN3 := #stringSecond, IN4 := 'S', IN5 := #stringMilliSecond, IN6 := 'MS');
   END_IF;

   IF (#tempDivHours > 0)
   THEN
     #tempStringTime := CONCAT(IN1 := #stringHour, IN2 := 'H', IN3 := #stringMinute, IN4 := 'M', IN5 := #stringSecond, IN6 := 'S', IN7 := #stringMilliSecond, IN8 := 'MS');
   END_IF;

   IF (#tempDivDays > 0)
   THEN
     #tempStringTime := CONCAT(IN1 := #stringDay, IN2 := 'D', IN3 := #stringHour, IN4 := 'H', IN5 := #stringMinute, IN6 := 'M', IN7 := #stringSecond, IN8 := 'S', IN9 := #stringMilliSecond, IN10 := 'MS');
   END_IF;

   // Write outputs
   #LGF_TimeToString := #tempStringTime;
END_FUNCTION

FUNCTION "LGF_BitsToWord" : Word   // FC10044, SCL
{ S7_Optimized_Access := 'TRUE' }
VERSION : 0.1
   VAR_INPUT
      bit0 : Bool;
      bit1 : Bool;
      bit2 : Bool;
      bit3 : Bool;
      bit4 : Bool;
      bit5 : Bool;
      bit6 : Bool;
      bit7 : Bool;
      bit8 : Bool;
      bit9 : Bool;
      bit10 : Bool;
      bit11 : Bool;
      bit12 : Bool;
      bit13 : Bool;
      bit14 : Bool;
      bit15 : Bool;
   END_VAR
BEGIN
   //=============================================================================
   // SIEMENS AG
   // (c)Copyright 2017
   //-----------------------------------------------------------------------------
   // Library:       LGF(Library General Functions)
   // Tested with:   CPU1212C DC/DC/DC FW:V4.2
   // Engineering:   TIA Portal V14 Update 1
   // Restrictions:  -
   // Requirements:  PLC (S7-1200 / S7-1500)
   // Functionality: This function converts 16 bits to a word
   //-----------------------------------------------------------------------------
   // Change log table:
   // Version  Date        In charge / Changes applied
   // 01.00.00 09.02.2017  Siemens Industry Online Support
   //                      First released version
   // 01.00.01 17.08.2018  Siemens Industry Online Support
   //                      Upgrade: TIA V15 Update 2
   // 01.00.02 23.11.2018  Siemens Industry Online Support
   //                      Upgrade: TIA V15.1
   //=============================================================================

   #LGF_BitsToWord.%X0 := #bit0;
   #LGF_BitsToWord.%X1 := #bit1;
   #LGF_BitsToWord.%X2 := #bit2;
   #LGF_BitsToWord.%X3 := #bit3;
   #LGF_BitsToWord.%X4 := #bit4;
   #LGF_BitsToWord.%X5 := #bit5;
   #LGF_BitsToWord.%X6 := #bit6;
   #LGF_BitsToWord.%X7 := #bit7;
   #LGF_BitsToWord.%X8 := #bit8;
   #LGF_BitsToWord.%X9 := #bit9;
   #LGF_BitsToWord.%X10 := #bit10;
   #LGF_BitsToWord.%X11 := #bit11;
   #LGF_BitsToWord.%X12 := #bit12;
   #LGF_BitsToWord.%X13 := #bit13;
   #LGF_BitsToWord.%X14 := #bit14;
   #LGF_BitsToWord.%X15 := #bit15;
END_FUNCTION

FUNCTION "LGF_WordToBits" : Void   // FC10045, SCL
{ S7_Optimized_Access := 'TRUE' }
VERSION : 0.1
   VAR_INPUT
      "word" : Word;
   END_VAR
   VAR_OUTPUT
      bit0 : Bool;
      bit1 : Bool;
      bit2 : Bool;
      bit3 : Bool;
      bit4 : Bool;
      bit5 : Bool;
      bit6 : Bool;
      bit7 : Bool;
      bit8 : Bool;
      bit9 : Bool;
      bit10 : Bool;
      bit11 : Bool;
      bit12 : Bool;
      bit13 : Bool;
      bit14 : Bool;
      bit15 : Bool;
   END_VAR
BEGIN
   //=============================================================================
   // SIEMENS AG
   // (c)Copyright 2017
   //-----------------------------------------------------------------------------
   // Library:       LGF(Library General Functions)
   // Tested with:   CPU1212C DC/DC/DC FW:V4.2
   // Engineering:   TIA Portal V14 Update 1
   // Restrictions:  -
   // Requirements:  PLC (S7-1200 / S7-1500)
   // Functionality: This function converts a word to 16 bits
   //-----------------------------------------------------------------------------
   // Change log table:
   // Version  Date        In charge / Changes applied
   // 01.00.00 09.02.2017  Siemens Industry Online Support
   //                      First released version
   // 01.00.01 17.08.2018  Siemens Industry Online Support
   //                      Upgrade: TIA V15 Update 2
   // 01.00.02 23.11.2018  Siemens Industry Online Support
   //                      Upgrade: TIA V15.1
   //=============================================================================

   #bit0 := #word.%X0;
   #bit1 := #word.%X1;
   #bit2 := #word.%X2;
   #bit3 := #word.%X3;
   #bit4 := #word.%X4;
   #bit5 := #word.%X5;
   #bit6 := #word.%X6;
   #bit7 := #word.%X7;
   #bit8 := #word.%X8;
   #bit9 := #word.%X9;
   #bit10 := #word.%X10;
   #bit11 := #word.%X11;
   #bit12 := #word.%X12;
   #bit13 := #word.%X13;
   #bit14 := #word.%X14;
   #bit15 := #word.%X15;
END_FUNCTION

